// TIA Portal project "ETI C 25" (V15.1)

(* hardware
DEVICE "ET 200SP station_1"  ET 200SP-Station
   slot 0: "Rack_0"  Rack  6ES5 710-8MAx1
   slot 1: "PLC_1"  CPU 1512SP-1 PN  6ES7 512-1DK01-0AB0  V2.6
   slot 2: "DI 16x24VDC ST_1"  DI 16x24VDC ST  6ES7 131-6BH01-0BA0  V0.0
      slot 1: "DI 16x24VDC ST_1"  DI 16x24VDC ST
   slot 3: "DI 16x24VDC ST_2"  DI 16x24VDC ST  6ES7 131-6BH01-0BA0  V0.0
      slot 1: "DI 16x24VDC ST_2"  DI 16x24VDC ST
   slot 4: "DQ 16x24VDC/0.5A ST_1"  DQ 16x24VDC/0.5A ST  6ES7 132-6BH01-0BA0  V0.0
      slot 1: "DQ 16x24VDC/0.5A ST_1"  DQ 16x24VDC/0.5A ST
   slot 5: "AQ 4xU/I ST_1"  AQ 4xU/I ST  6ES7 135-6HD00-0BA1  V1.1
      slot 1: "AQ 4xU/I ST_1"  AQ 4xU/I ST
   slot 6: "Server module_1"  Server module  6ES7 193-6PA00-0AA0  V1.1
      slot 1: "Server module_1"  Server module
   slot 127: "BA 2xRJ45"  BA 2xRJ45  6ES7 193-6AR00-0AA0  V0.0
      slot 32769: "Port_1"  6ES7 193-6AR00-0AA0
      slot 32770: "Port_2"  6ES7 193-6AR00-0AA0
DEVICE "GSD device_1"  GSD.Device.PN
   slot 0: "Rack"  Rack  V1.0
   slot 0: "IOL_I_16_HUB"  IOL_I/O_ 4/ 4 Byte
   slot 0: "mvk1"  55162 MVK DIO12 DIO4/IOL4 M12L 4P  55162  1.08.10
      slot 0: "55162 MVK DIO12 DIO4/IOL4 M12L 4P_1"  55162 MVK DIO12 DIO4/IOL4 M12L 4P
      slot 1: "55162 MVK DIO12 DIO4/IOL4 M12L 4P 1"  55162 MVK DIO12 DIO4/IOL4 M12L 4P
         slot 1: "Port 1"  Port 1
         slot 2: "Port 2"  Port 2
      slot 1: "Device_1"  Device
         slot 0: "Parameter/Diagnostic"  Parameter/Diagnostic
         slot 1: "Digital IO"  Digital IO
      slot 2: "IO-Link master_1"  IO-Link master
   slot 1: "Deactivated"  Deactivated
   slot 2: "Qualifier DI"  Qualifier DI
   slot 2: "FESTO_propocionalniVentil"  IOL_I/O_ 8/ 8 Byte
   slot 3: "Qualifier DO"  Qualifier DO
   slot 3: "SDAT1"  IOL_I_ 2 Byte
   slot 4: "System state"  System state
DEVICE "GSD device_2"  GSD.Device.PN
   slot 0: "Rack"  Rack  V1.0
   slot 0: "IOL_I/O_ 4/ 4 Byte"  IOL_I/O_ 4/ 4 Byte
   slot 0: "mvk2"  55162 MVK DIO12 DIO4/IOL4 M12L 4P  55162  1.08.10
      slot 0: "55162 MVK DIO12 DIO4/IOL4 M12L 4P_1"  55162 MVK DIO12 DIO4/IOL4 M12L 4P
      slot 1: "55162 MVK DIO12 DIO4/IOL4 M12L 4P 2"  55162 MVK DIO12 DIO4/IOL4 M12L 4P
         slot 1: "Port 1"  Port 1
         slot 2: "Port 2"  Port 2
      slot 1: "Device_1"  Device
         slot 0: "Parameter/Diagnostic"  Parameter/Diagnostic
         slot 1: "Digital IO"  Digital IO
      slot 2: "IO-Link master_1"  IO-Link master
   slot 1: "MURR_MVP_2"  IOL_I_ 2 Byte
   slot 2: "Qualifier DI"  Qualifier DI
   slot 2: "IOL_BANNER_LED"  IOL_O_ 4 Byte
   slot 3: "Qualifier DO"  Qualifier DO
   slot 3: "FESTO_SDE1_PRITISK"  IOL_I_ 2 Byte
   slot 4: "System state"  System state
DEVICE "GSD device_3"  GSD.Device.PN
   slot 0: "Rack"  Rack  V1.0
   slot 0: "mvk3"  54504 SOLID67 IOL8 60mm M12L 5P  54504  2.1.1
      slot 0: "DAP"  DAP
      slot 1: "PN-IO"  PN-IO
         slot 1: "Port X01 10/100 MBit/s"  Port X01 10/100 MBit/s
         slot 2: "Port X02 10/100 MBit/s"  Port X02 10/100 MBit/s
      slot 1: "IO-Link Master_1"  IO-Link Master  1.0
         slot 0: "Status/Control Module"  Status/Control Module  1.0
   slot 1: "IFM_VS_temp_pretok"  IO-Link In 4 Bytes
   slot 2: "Digital In (A)/Dig. (B)_1"  Digital In (A)/Dig. (B)
   slot 3: "Digital In (A)/Dig. (B)_2"  Digital In (A)/Dig. (B)
   slot 4: "Digital In (A)/Dig. (B)_3"  Digital In (A)/Dig. (B)
   slot 5: "Digital Out (A)/Dig. (B)"  Digital Out (A)/Dig. (B)
   slot 6: "Digital Out (A)/Dig. (B)_1"  Digital Out (A)/Dig. (B)
   slot 7: "Kamera"  Digital In (A)/Dig. (B)
   slot 8: "FESTO Pnevmatski BLok IO-Link I/O 8/8 Bytes"  IO-Link I/O 8/8 Bytes
DEVICE "GSD device_4"  GSD.Device.PN
   slot 0: "Rack"  Rack  V1.0
   slot 0: "varilnik"  PSS6000 Weld Timer (2-Port)  PSS6000  V1.13.1
      slot 0: "RT"  RT
      slot 1: "Interface"  Interface
         slot 1: "Port 1"  Port 1
         slot 2: "Port 2"  Port 2
   slot 1: "PSI6xxx.780_1"  PSI6xxx.780
      slot 0: "PSI6xxx.780"  PSI6xxx.780
DEVICE "GSD device_7"  GSD.Device.PN
   slot 0: "Rack"  Rack  V1.0
   slot 0: "akd"  AKD-PN-DEVICE  AKD-Pxxxxx-xxPN-xxxx  V00.02
      slot 0: "IDS_SUBMODULE_PARAMDAP"  IDS_SUBMODULE_PARAMDAP
      slot 1: "Interface"  Interface
         slot 1: "Port_1"  Port
   slot 1: "Standard telegram 9_1"  Standard telegram 9  1.0
      slot 0: "Standard telegram 9"  Standard telegram 9
DEVICE "GSD device_5"  GSD.Device.PN
   slot 0: "Rack"  Rack  V1.0
   slot 0: "kroznik"  AKD-PN-DEVICE  AKD-Pxxxxx-xxPN-xxxx  V00.02
      slot 0: "IDS_SUBMODULE_PARAMDAP"  IDS_SUBMODULE_PARAMDAP
      slot 1: "Interface"  Interface
         slot 1: "Port_1"  Port
   slot 1: "Standard telegram 9_1"  Standard telegram 9  1.0
      slot 0: "Standard telegram 9"  Standard telegram 9
DEVICE "GSD device_6"  GSD.Device.PN
   slot 0: "Rack"  Rack  V1.0
   slot 0: "cilinder"  AKD-PN-DEVICE  AKD-Pxxxxx-xxPN-xxxx  V00.02
      slot 0: "IDS_SUBMODULE_PARAMDAP"  IDS_SUBMODULE_PARAMDAP
      slot 1: "Interface"  Interface
         slot 1: "Port_1"  Port
   slot 1: "Standard telegram 9_1"  Standard telegram 9  1.0
      slot 0: "Standard telegram 9"  Standard telegram 9
DEVICE "TP1200 Comfort"  TP1200 Comfort
   slot 0: "TP1200 Comfort"  TP1200 Comfort  6AV2 124-0MC01-0AX0  15.0.0.0
   slot 1: "HMI_RT_6"  TP1200 Comfort  6AV2 124-0MC01-0AX0  15.0.0.0
   slot 5: "TP900 Comfort._CP_1"  PROFINET Interface  15.0.0.0
      slot 1: "PROFINET Interface_1"  PROFINET Interface
         slot 1: "Port_1"  Port
         slot 2: "Port_2"  Port
   slot 7: "TP900 Comfort.I/DP_CP_1"  MPI/DP Interface  15.0.0.0
DEVICE "GSD device_8"  GSD.Device.PN
   slot 0: "Rack"  Rack  V1.0
   slot 0: "dl-pn1"  DL-PN1  DL-PN1  1.00
      slot 0: "DL-PN1"  DL-PN1  1.00
      slot 1: "Interface"  Interface
         slot 1: "Port 1"  Port 1
   slot 1: "DL-PN1_1"  DL-PN1
      slot 0: "DL-PN1 Device"  DL-PN1 Device
   slot 2: "GT2-***_1"  GT2-***
      slot 0: "GT2-***"  GT2-***
   slot 3: "GT2-***_2"  GT2-***
      slot 0: "GT2-***"  GT2-***
*)

// ===== PLC "PLC_1"  CPU 1512SP-1 PN =====

VAR_GLOBAL   // PLC tag table "Default tag table"
   "System_Byte" AT %MB1 : Byte;
   "FirstScan" AT %M1.0 : Bool;
   "DiagStatusUpdate" AT %M1.1 : Bool;
   "AlwaysTRUE" AT %M1.2 : Bool;
   "AlwaysFALSE" AT %M1.3 : Bool;
   "Clock_Byte" AT %MB0 : Byte;
   "Clock_10Hz" AT %M0.0 : Bool;
   "Clock_5Hz" AT %M0.1 : Bool;
   "Clock_2.5Hz" AT %M0.2 : Bool;
   "Clock_2Hz" AT %M0.3 : Bool;
   "Clock_1.25Hz" AT %M0.4 : Bool;
   "Clock_1Hz" AT %M0.5 : Bool;
   "Clock_0.625Hz" AT %M0.6 : Bool;
   "Clock_0.5Hz" AT %M0.7 : Bool;
   "Tag_1" AT %M20.0 : Bool;
   "Tag_2" AT %QD24 : DWord;
   "Tag_3" AT %MD400 : DWord;
   "Tag_4" AT %QD28 : DWord;
   "STOP_SR" AT %M2.0 : Bool;
   "RočnoMerker" AT %M2.2 : Bool;
   "vkloprocno" AT %M2.6 : Bool;
   "RežimDelovanja" AT %MB3 : Byte;
   "BANNER_B3" AT %QB25 : Byte;
   "BANNER_B2" AT %QB26 : Byte;
   "BANNER_B1" AT %QB27 : Byte;
   "BANNER_B0" AT %QB28 : Byte;
   "Tag_5" AT %QW28 : Word;
   "Tag_6" AT %QW25 : Word;
   "Tag_7" AT %QD25 : DWord;
   "STEVEC_KONEC_TRAKA_DOSEZEN" AT %M4.1 : Bool;
   "StatusPrisotnostiTraku" AT %MB5 : Byte;
   "NapakaOdvijanjaTrau" AT %M4.2 : Bool;   // Napaka če se srebrn trak ne odvije
   "NapakaCiscenjaElektrode" AT %M4.3 : Bool;   // Napaka Motorja Čiščenja Traku
   "CiscenjeElektrodeManualOn" AT %M4.4 : Bool;
   "RocniVKlopOdvijanjaTraku" AT %M4.5 : Bool;
   "IzklopStroja" AT %M4.6 : Bool;
   "stevecpreklopov" AT %ID4 : DInt;
   "ZavarjenoSlabiKosi" AT %MD6 : DInt;
   "StartUpBit" AT %M4.7 : Bool;
   "kameratrigger" AT %M10.0 : Bool;
   "ST_IZDELKOV" AT %MD16 : DInt;   // STEVEC KOSOV
END_VAR

VAR_GLOBAL   // PLC tag table "MVK1"
   "MVK_b0" AT %IB20 : Byte;
   "MVK_b1" AT %IB21 : Byte;
   "MVK_b2" AT %IB22 : Byte;
   "MVK_b3" AT %IB23 : Byte;
   "MVK_dw" AT %ID20 : DWord;
   "MVK1_w0" AT %IW20 : Word;
   "ZaporaIzdelka" AT %I20.0 : Bool;   // Y1/1
   "SprositevZaporeIzdelka" AT %I20.1 : Bool;   // Y1/1
   "PrijemaloKontaktaZaprto" AT %I20.2 : Bool;   // Y3/1
   "PrijemaloKontaktaOdprto" AT %I20.3 : Bool;   // Y3/1
   "PozKontaktNaKoncuLetve" AT %I20.4 : Bool;   // Kontakt na koncu letve
   "NC_20.5" AT %I20.5 : Bool;   // NC
   "PozKontaktNaprej" AT %I20.6 : Bool;   // Pozicioniranje pred varjenjem
   "PozKontaktNazaj" AT %I20.7 : Bool;   // Pozicioniranjem pred varjenjem
   "DrzanjeIzmetKontakta" AT %I21.0 : Bool;   // Odpiranje dzanja kontakta nazaj
   "DrzanjeKontakta" AT %I21.1 : Bool;   // Izmet kontakta nazaj
   "IzmetKontaktaNazaj" AT %I21.2 : Bool;   // Izmet vzvoda je v izhodiscu
   "NC_21.3" AT %I21.3 : Bool;   // NC
   "DrcaDobriKosi" AT %I21.4 : Bool;   // Pozicija za dobre kose
   "DrscaSLabiKosi" AT %I21.5 : Bool;   // Pozicija za slabe kose
   "SenzorOdvijanjaCiscenjeElektrode" AT %I21.6 : Bool;   // SenzorCiscenjaElektrode
   "NC_21.7" AT %I21.7 : Bool;
END_VAR

VAR_GLOBAL   // PLC tag table "MVK2"
   "MVK2_b0" AT %IB8 : Byte;
   "MVK2_b1" AT %IB9 : Byte;
   "MVK2_b2" AT %IB10 : Byte;
   "MVK2_b3" AT %IB11 : Byte;
   "MVK2_dw" AT %ID8 : DWord;
   "MVK2_w0" AT %IW8 : Word;
   "MVK2_w1" AT %IW10 : Word;
   "KAMERA_FEEDBACK" AT %I8.0 : Bool;
   "NC_8.1" AT %I8.1 : Bool;
   "NC_8.2" AT %I8.2 : Bool;
   "NC_8.3" AT %I8.3 : Bool;
   "SenzorStartOdvijanje" AT %I8.4 : Bool;   // Senzor za začetek odvijanja koluta
   "SenzorKoluta" AT %I8.5 : Bool;   // Senzor za detekcijo odvijanja koluta
   "PrisotnostTraka" AT %I8.6 : Bool;
   "NC_8.7" AT %I8.7 : Bool;
   "RazsvetljavaLevo" AT %Q20.0 : Bool;
   "RazsvetljavaDesno" AT %Q20.1 : Bool;
   "NC_Q20.2" AT %Q20.2 : Bool;
   "NC_Q20.3" AT %Q20.3 : Bool;
   "NC_Q20.4" AT %Q20.4 : Bool;
   "NC_Q20.5" AT %Q20.5 : Bool;
   "NC_Q20.6" AT %Q20.6 : Bool;
   "NC_Q20.7" AT %Q20.7 : Bool;
END_VAR

VAR_GLOBAL   // PLC tag table "SDAT"
   "I_SDAT1" AT %IW32 : Word;   // Y2/1
   "I_SDAT2" AT %IW34 : Word;   // Y1/2
END_VAR

VAR_GLOBAL   // PLC tag table "MURR IOL M"
   "MURR_IOL1_DO" AT %QB0 : Byte;
   "SoftStart" AT %Q0.0 : Bool;   // SOFTSTART - vklop pnevmatike
   "MURR_IOL1_DO.1" AT %Q0.1 : Bool;
   "MURR_IOL1_DO.2" AT %Q0.2 : Bool;   // Napajanje IOL power supply
   "MURR_IOL1_DO.3" AT %Q0.3 : Bool;
   "MURR_IOL1_DO.4" AT %Q0.4 : Bool;
   "MURR_IOL1_DO.5" AT %Q0.5 : Bool;
   "MURR_IOL1_DO.6" AT %Q0.6 : Bool;
   "MURR_IOL1_DO.7" AT %Q0.7 : Bool;
   "MURR_IOL2_DO" AT %QB2 : Byte;
   "MURR_IOL2_DO.0" AT %Q2.0 : Bool;
   "MURR_IOL2_DO.1" AT %Q2.1 : Bool;
   "MURR_IOL2_DO.2" AT %Q2.2 : Bool;
   "MURR_IOL2_DO.3" AT %Q2.3 : Bool;
   "MURR_IOL2_DO.4" AT %Q2.4 : Bool;
   "MURR_IOL2_DO.5" AT %Q2.5 : Bool;
   "MURR_IOL2_DO.6" AT %Q2.6 : Bool;
   "MURR_IOL2_DO.7" AT %Q2.7 : Bool;
   "FESTO_pritisk" AT %IW52 : Word;
   "PropocionalniVentilSet" AT %QW32 : Word;
   "PropocionalniVentilTrenutna" AT %IW44 : Word;
END_VAR

VAR_GLOBAL   // PLC tag table "FESTO"
   "FESTO_W0" AT %QW44 : Word;
   "FESTO_W1" AT %QW46 : Word;
   "FESTO_W2" AT %QW48 : Word;
   "FESTO_W3" AT %QW50 : Word;
   "1Y1_OdklepZapore" AT %Q44.0 : Bool;
   "Y2/1_NalaganjeNaprej" AT %Q44.2 : Bool;
   "Y2/1_NalaganjeNazanj" AT %Q44.3 : Bool;
   "Y3/1_PrijemaloKontaktaOdpri" AT %Q44.4 : Bool;
   "Y3/1_NC" AT %Q44.5 : Bool;
   "Y1/3_OdmičniCilinderKonusa" AT %Q45.0 : Bool;
   "Y1/3_NC" AT %Q45.1 : Bool;
   "Y2/3_PozicioniranjeKontaktovNazaj" AT %Q45.2 : Bool;
   "Y2/3_PozicioniranjeKontaktovNaprej" AT %Q45.3 : Bool;
   "Y3/3_OdpiranjeDržalaKomada" AT %Q45.4 : Bool;
   "Y3/3_NC" AT %Q45.5 : Bool;
   "Y4/3_OdpiranjeIzmetaKontakta" AT %Q45.6 : Bool;
   "Y4/3_NC" AT %Q45.7 : Bool;
   "Y5/3_IzmetKomadov" AT %Q46.0 : Bool;
   "Y5/3_NC" AT %Q46.1 : Bool;
   "Y6/3_LoputaDobri" AT %Q46.2 : Bool;
   "Y6/3_LoputaSlabi" AT %Q46.3 : Bool;
   "Y1/4_odmičniCilinderVarjenje_GOR" AT %Q46.4 : Bool;
   "Y1/4_odmičniCilinderVarjenjeDOL" AT %Q46.5 : Bool;
   "ČiščenjeElektrode_ON" AT %Q46.6 : Bool;
   "ČiščenjeElektrode_OFF" AT %Q46.7 : Bool;
   "PihanjeLinearniVibrator" AT %Q47.0 : Bool;
   "NC" AT %Q47.1 : Bool;
   "Y2/1_dovajanjePlosciceNazaj" AT %Q44.6 : Bool;
   "Y2_1_dovajanjePlosciceNaprej" AT %Q44.7 : Bool;
   "1Y1_zaklep_NC" AT %Q44.1 : Bool;
END_VAR

VAR_GLOBAL   // PLC tag table "MVK3"
   "MVK3_b0" AT %QB40 : Byte;
   "MVK3_b1" AT %QB41 : Byte;
   "MVK3_b2" AT %QB42 : Byte;
   "MVK3_b4" AT %QB43 : Byte;
   "MVK3_O_X1_P4" AT %Q40.0 : Bool;
   "MVK3_O_X1_P2" AT %Q40.1 : Bool;
   "MVK3_O_X2_P4" AT %Q40.2 : Bool;
   "MVK3_O_X2_P2" AT %Q40.3 : Bool;
   "MVK3_O_X3_P4" AT %Q40.4 : Bool;
   "MVK3_O_X3_P2" AT %Q40.5 : Bool;
   "MVK3_O_X4_P4" AT %Q40.6 : Bool;
   "MVK3_O_X4_P2" AT %Q40.7 : Bool;
   "MVK3_O_X5_P4_NC" AT %Q41.0 : Bool;   // X5,P4 - PIN 4 NC
   "RazsvetljavaSpredaj" AT %Q41.1 : Bool;   // 5404 IOL X5, P2 - MASTER - PIN2/5 - razsvetljava LED SPREDAJ
   "bTrigOptoEnginering" AT %Q41.2 : Bool;   // X6, P4 : triger za led
   "bVccOptoEngineering" AT %Q41.3 : Bool;   // X6, P2 : Vklop napajanja
   "MVK3_O_b1.4" AT %Q41.4 : Bool;   // X7, P4
   "MVK3_O_b1.5" AT %Q41.5 : Bool;   // X7, P2
   "MVK3_O_b1.6" AT %Q41.6 : Bool;   // X8, P4
   "MVK3_O_b1.7" AT %Q41.7 : Bool;   // X8,P2
   "MVK3_O_b2.0" AT %Q42.0 : Bool;
   "MVK3_O_b2.1" AT %Q42.1 : Bool;
   "MVK3_O_b2.2" AT %Q42.2 : Bool;
   "MVK3_O_b2.3" AT %Q42.3 : Bool;
   "MVK3_O_b2.4" AT %Q42.4 : Bool;
   "MVK3_O_b2.5" AT %Q42.5 : Bool;
   "MVK3_O_b2.6" AT %Q42.6 : Bool;
   "MVK3_O_b2.7" AT %Q42.7 : Bool;
   "MVK3_O_b3.0" AT %Q43.0 : Bool;
   "MVK3_O_b3.1" AT %Q43.1 : Bool;
   "MVK3_O_b3.2" AT %Q43.2 : Bool;
   "MVK3_O_b3.3" AT %Q43.3 : Bool;
   "MVK3_O_b3.4" AT %Q43.4 : Bool;
   "MVK3_O_b3.5" AT %Q43.5 : Bool;
   "MVK3_O_b3.6" AT %Q43.6 : Bool;
   "MVK3_O_b3.7" AT %Q43.7 : Bool;
   "IOL_IFM_SV" AT %ID36 : DWord;
   "MVK3_I_b0" AT %IB54 : Byte;
   "MVK3_I_b1" AT %IB55 : Byte;
   "MVK3_I_b2" AT %IB56 : Byte;
   "MVK3_I_b3" AT %IB57 : Byte;
END_VAR

VAR_GLOBAL   // PLC tag table "PLC_IO"
   "PLC_I_W0" AT %IW0 : Word;
   "PLCI_W2" AT %IW2 : Word;
   "PLC_I0.0" AT %I0.0 : Bool;   // DC OK
   "IzklopVsiliBtnPanel" AT %I0.1 : Bool;
   "VarmostZavese" AT %I0.2 : Bool;   // VarnostneZavese [1-ok, 0, nok]
   "PremostitevVarnostiBtnPanel" AT %I0.3 : Bool;
   "PrisotnostIzmetaIzdelka" AT %I0.4 : Bool;   // Senzor Izmeta na koncu traku
   "PLC_I0.5" AT %I0.5 : Bool;
   "PLC_I0.6" AT %I0.6 : Bool;
   "PLC_I0.7" AT %I0.7 : Bool;
   "PLC_I1.0" AT %I1.0 : Bool;
   "PLC_I1.1" AT %I1.1 : Bool;
   "RežimRočno" AT %I1.2 : Bool;
   "RežimAvtomatsko" AT %I1.3 : Bool;
   "StartCiklaBtnPanel" AT %I1.4 : Bool;
   "StopCiklaBtnPanel" AT %I1.5 : Bool;
   "ResetNapake" AT %I1.6 : Bool;
   "VklopKrmiljaBtnPanel" AT %I1.7 : Bool;
   "VKlopvarnostnegaModulaIVS" AT %QW4 : Word;
   "VklopVarnosnegaModula" AT %Q4.0 : Bool;
   "VklopZaves" AT %Q4.1 : Bool;
   "NightShift" AT %Q4.2 : Bool;
   "AKD_sprostitevZavore" AT %Q4.3 : Bool;
   "PLC_Q4.4" AT %Q4.4 : Bool;
   "PLC_Q4.5" AT %Q4.5 : Bool;
   "PLC_Q4.6" AT %Q4.6 : Bool;
   "VentilVode" AT %Q4.7 : Bool;
   "PLC_Q5.0" AT %Q5.0 : Bool;
   "MotorOdvijanjeTraku" AT %Q5.1 : Bool;
   "MotorČiščenjeElektrode" AT %Q5.2 : Bool;
   "LED_RUN" AT %Q5.3 : Bool;
   "LED_ERROR" AT %Q5.4 : Bool;
   "AKD_HW_ENABLE" AT %Q5.5 : Bool;
   "TekociTrakVklop" AT %Q5.6 : Bool;
   "PolnjenjeSkatle1" AT %Q5.7 : Bool;
   "+" AT %I2.0 : Bool;
   "-" AT %I2.1 : Bool;
   "i2.0_b2" AT %I2.2 : Bool;
   "i2.0_b3" AT %I2.3 : Bool;
   "i2.0_b4" AT %I2.4 : Bool;
   "i2.0_b5" AT %I2.5 : Bool;
   "i2.0_b6" AT %I2.6 : Bool;
   "i2.0_b7" AT %I2.7 : Bool;
   "i2.0_b8" AT %I3.0 : Bool;
   "i2.0_b9" AT %I3.1 : Bool;
   "i2.0_b10" AT %I3.2 : Bool;
   "i2.0_b11" AT %I3.3 : Bool;
   "i2.0_b12" AT %I3.4 : Bool;
   "i2.0_b13" AT %I3.5 : Bool;
   "i2.0_b14" AT %I3.6 : Bool;
END_VAR

VAR_GLOBAL   // PLC tag table "VARJENJE"
   "Varjenje_QB0" AT %QB52 : Byte;
   "Varjenje_QB1" AT %QB53 : Byte;
   "Varjanje_IB0" AT %IB66 : Byte;
   "Varjenje_IB0" AT %IB67 : Byte;
   "ValidSpotSelection" AT %Q52.0 : Bool;
   "Varjenje_Qb0.1" AT %Q52.1 : Bool;
   "Start" AT %Q52.2 : Bool;
   "GeneralFaultReset" AT %Q52.3 : Bool;
   "ResetWithEOS" AT %Q52.4 : Bool;
   "ResetWithReweld" AT %Q52.5 : Bool;
   "Varjenje_Qb0.6" AT %Q52.6 : Bool;
   "Varjenje_Qb0.7" AT %Q52.7 : Bool;
   "ExternalWeldOn" AT %Q53.0 : Bool;
   "Varjenje_Qb1.1" AT %Q53.1 : Bool;
   "Varjenje_Qb1.2" AT %Q53.2 : Bool;
   "Varjenje_Qb1.3" AT %Q53.3 : Bool;
   "Varjenje_Qb1.4" AT %Q53.4 : Bool;
   "Varjenje_Qb1.5" AT %Q53.5 : Bool;
   "Varjenje_Qb1.6" AT %Q53.6 : Bool;
   "Varjenje_Qb1.7" AT %Q53.7 : Bool;
   "Varjenje_Qb2.0" AT %Q54.0 : Bool;
   "Varjenje_Qb2.1" AT %Q54.1 : Bool;
   "Varjenje_Qb2.2" AT %Q54.2 : Bool;
   "Varjenje_Qb2.3" AT %Q54.3 : Bool;
   "Varjenje_Qb2.4" AT %Q54.4 : Bool;
   "Varjenje_Qb2.5" AT %Q54.5 : Bool;
   "Varjenje_Qb2.7" AT %Q54.7 : Bool;
   "Varjenje_Qb2.8" AT %Q55.0 : Bool;
   "Varjenje_Qb2.9" AT %Q55.1 : Bool;
   "Varjenje_Qb2.10" AT %Q55.2 : Bool;
   "Varjenje_Qb2.11" AT %Q55.3 : Bool;
   "Varjenje_Qb2.12" AT %Q55.4 : Bool;
   "SpotSelection" AT %QB60 : Byte;
   "SpotSelectionTakeOver" AT %I66.0 : Bool;   // Program izbran
   "Varjenje_Ib0.1" AT %I66.1 : Bool;
   "EndOfSequency_WC" AT %I66.2 : Bool;   // Konec varjenja
   "TimerReady" AT %I66.3 : Bool;   // Varilnik pripravljen
   "WeldFault" AT %I66.4 : Bool;   // Napaka varjenja
   "Varjenje_Ib0.5" AT %I66.5 : Bool;
   "Varjenje_Ib0.6" AT %I66.6 : Bool;
   "Varjenje_Ib0.7" AT %I66.7 : Bool;
   "FiringEnable" AT %I67.0 : Bool;   // Varjenje Vključeno
   "Varjenje_Ib2.1" AT %I67.1 : Bool;
   "Varjenje_Ib2.2" AT %I67.2 : Bool;
   "Varjenje_Ib2.3" AT %I67.3 : Bool;
   "Varjenje_Ib2.4" AT %I67.4 : Bool;
   "Varjenje_Ib2.5" AT %I68.0 : Bool;
   "Varjenje_Ib2.6" AT %I68.1 : Bool;
   "Varjenje_Ib2.7" AT %I68.2 : Bool;
   "Varjenje_Ib2.8" AT %I68.3 : Bool;
   "Varjenje_Ib2.9" AT %I68.4 : Bool;
   "Varjenje_Ib2.10" AT %I68.5 : Bool;
   "StatusCode" AT %IB82 : Byte;   // Status
   "Status_b0" AT %IB80 : Byte;
   "Status_b1" AT %IB83 : Byte;
   "Varjenje_Qb2.6" AT %Q54.6 : Bool;
END_VAR

VAR_GLOBAL   // PLC tag table "AKD_elektroda"
   "PogojZaservoOn" AT %M2.1 : Bool;
   "tipka+" AT %M2.3 : Bool;
   "tipka-" AT %M2.4 : Bool;
   "ElektrodaSiemensToAkd" AT %Q400.0 : "SIEMENS_TO_AKD";
   "ElektrodaAkdToSiemens" AT %I400.0 : "AKD_TO_SIEMENS";
   "onemogoci" AT %M2.7 : Bool;
   "enable" AT %M4.0 : Bool;
   "STEVEC_KOSOV" AT %C0 : Counter;
   "manualCameraTrig" AT %M10.1 : Bool;   // trig kamera
   "MotorCiscenjeElektrodeCOunter" AT %MD12 : DInt;   // Stevec
   "prisotnostizmetaarker" AT %M10.2 : Bool;   // Merker za R edge - izmeta kontakta - senzor
END_VAR

VAR_GLOBAL   // PLC tag table "AKD_kroznik"
   "KroznikSiemensToAkd" AT %Q98.0 : "SIEMENS_TO_AKD";
   "KroznikAkdToSiemens" AT %I98.0 : "AKD_TO_SIEMENS";
   "servpen" AT %M2.5 : Bool;
END_VAR

VAR_GLOBAL   // PLC tag table "AKD_REZANJEPODAJANJE"
   "rezanjepodajanjeSiemenstoAKD" AT %I108.0 : "AKD_TO_SIEMENS";
   "rezanjepodajanje_SiemensToAKD" AT %Q118.0 : "SIEMENS_TO_AKD";
END_VAR

VAR_GLOBAL   // PLC tag table "KEYENCE"
   "Keyence_OdmičniCilinderKonusa" AT %ID137 : DInt;   // Cilinder odmika mize
   "Keyence_OdmičniCilinderVarjenja" AT %ID144 : DInt;   // Cilinder odmika varjenja
END_VAR

TYPE "UDT_MVK1"
   STRUCT
      "1Y1" : Struct   // VKLOP/IZKLOP zapore na LIN vibratorju
         B1 : Bool;   // POZ Zaklep linearnega vibratorja
         B2 : Bool;   // POZ Odklep linearnega vibratorja
      END_STRUCT;
      "Y3/1" : Struct   // Prijemalo kontakta
         B1 : Bool;   // POZ Prijemalo zaprto
         B2 : Bool;   // POZ Prijemalo odprto
      END_STRUCT;
      B_kontaktnaKoncuLetve : Struct   // Detekcija kontakta na letvi
         B1 : Bool;   // POZ kontakt na koncu letve
         NC : Bool;
      END_STRUCT;
      "Y2/3" : Struct   // Pozicioniranje kontakta
         B1 : Bool;   // POZ kontakta naprej
         B2 : Bool;   // POZ Prijemalo odprto
      END_STRUCT;
      "Y3/3" : Struct   // Držanje kontakta v mizi
         B1 : Bool;   // POZ držanje kontakta odprto
      END_STRUCT;
      "Y4/3" : Struct   // Odpiranje izmeta konkta
         B1 : Bool;   // POZ izmet kontakta odprt
      END_STRUCT;
      "Y5/3" : Struct   // Izmet kontakta
         B1 : Bool;   // POZ izmet kontakta nazaj
      END_STRUCT;
      "Y6/3" : Struct   // Drča dobri/slabi kosi
         B1 : Bool;   // POZ dobri kosi
         B2 : Bool;   // POZ slabi kosi
      END_STRUCT;
      KonrolaIzmeta : Struct   // kontrola izmeta
         IzmetOK : Bool;   // Senzor preleta izmeta
         NC : Bool;
      END_STRUCT;
   END_STRUCT;
END_TYPE

TYPE "SIEMENS_TO_AKD"
   STRUCT
      PODATKI : Struct
         oBit8_jogOn : Bool;   // b0
         oBit9_jog2On : Bool;   // 1
         ControlByPLC : Bool;   // 2
         StartHomming : Bool;   // 3
         NC_B0_b4 : Bool;   // 4
         NC_B0_b5 : Bool;   // 5
         NC_B0_b6 : Bool;   // 6
         NC_B0_b7 : Bool;   // 7
         SwtichOn : Bool;   // 0
         NoCoastStop : Bool;   // 1
         NoQuickStop : Bool;   // 2
         EnableOperation : Bool;   // 3
         EnableRampGen : Bool;   // 4
         UnfreezeRamp : Bool;   // 5
         EnableSetPoint : Bool;   // 6
         FaultAckt : Bool;   // 7 1
         SATANW : Int;   // 0- 26 2-3
         byte4 : Byte;   // 4
         byte5 : Byte;   // 5
         MDI_TARPOS : DInt;   // 6 7 8 9
         MDI_VELOCITY : DInt;   // 10 11 12 13
         b14 : DInt;   // 14
         "15" : DInt;   // 15
         b16 : DInt;   // 16
         b17 : DInt;   // 17
         MDI_MOD : DInt;   // 18,19
      END_STRUCT;
   END_STRUCT;
END_TYPE

TYPE "AKD_TO_SIEMENS"
   STRUCT
      PODATKI_TO_SIEMENS : Struct
         ErrInRange : Bool;
         ContrReqByMass : Bool;
         TargetPosreached : Bool;
         HomePosSet : Bool;
         TravesingTaskAck : Bool;
         DriveStopen : Bool;
         MotionTaskActive : Bool;
         "i_b0.7" : Bool;
         ReadyToSwitch : Bool;
         ReadyToOperate : Bool;
         OperationENabled : Bool;
         FaultPresent : Bool;
         CoastStopNotAct : Bool;
         QuickStopNotAct : Bool;
         SwitchOnInhibiited : Bool;
         WarningPreent : Bool;
         AKTSATZ : Word;
         ZSW2 : Word;
         ActualPos : DWord;
      END_STRUCT;
   END_STRUCT;
END_TYPE

TYPE "PDT_AKD"
   STRUCT
      PODATKI : Struct
         AKDenable : Bool;
         NastavitevHitrosti : Int := 60;
         NastavitevPozicije : DInt := 12;
         TrenutnaPozicija : DInt;
         ServoGo : Bool;
         StartHomming : Bool;
      END_STRUCT;
   END_STRUCT;
END_TYPE

TYPE "BOSH"
   STRUCT
      PDT_BOSH_STATUS : Struct
         OK : UInt := 0;
         IZKLOP_V_SILI : UInt := 80;
         WELD_WITHOUD_COMMAND : UInt := 81;
         MEMMORY_DELETED : UInt := 85;
         DATA_DOWNLOAD_ACTIVE : UInt := 86;
         NO_WELDING_PROGRAM : UInt := 87;
         HARDWARE_FAULT : UInt := 88;
         "I/O_BUS_FAULT" : UInt := 89;
         HWAVE_MONITORING : UInt := 90;
         MAIN_SWITCH_TRIPPED : UInt := 91;
         EXTERNAL_TEMEPERATURE_TO_HIGH : UInt := 92;
         SYC_ERROR : UInt := 93;
         START_INHIBITED : UInt := 94;
         PROGRAM_PARITY_ERROR : UInt := 95;
         PROGRAMED_VALUE_TO_LARGE : UInt := 98;
         WELD_PROCESS_ERROR : UInt := 99;
         SUPPLY_VOLTAGE_VAULT : UInt := 100;
         MAX_HEAT_SINK_TEMP : UInt := 160;
         TRANSFORMER_TEMP_TO_HIGH : UInt := 164;
         HARDWARE_FAULT_DRIVE_MODULE : UInt := 165;
      END_STRUCT;
   END_STRUCT;
END_TYPE

DATA_BLOCK "SDAT1"   // DB1
{ S7_Optimized_Access := 'TRUE' }
VERSION : 0.1
// stored: InstanceOfName FB_IOL_SDAT
"FB_IOL_SDAT"
BEGIN
END_DATA_BLOCK

DATA_BLOCK "SDAT2"   // DB2
{ S7_Optimized_Access := 'TRUE' }
VERSION : 0.1
// stored: InstanceOfName FB_IOL_SDAT
"FB_IOL_SDAT"
BEGIN
END_DATA_BLOCK

DATA_BLOCK "FB_MVK1_DB"   // DB3
{ S7_Optimized_Access := 'TRUE' }
VERSION : 0.1
// stored: InstanceOfName FB_MVK1
"FB_MVK1"
BEGIN
END_DATA_BLOCK

DATA_BLOCK "FB_IOL_IFM_SV_DB"   // DB4
{ S7_Optimized_Access := 'TRUE' }
VERSION : 0.1
// stored: InstanceOfName FB_IOL_IFM_SV
"FB_IOL_IFM_SV"
BEGIN
END_DATA_BLOCK

DATA_BLOCK "FB_FESTO_VPPM_DB"   // DB5
{ S7_Optimized_Access := 'TRUE' }
VERSION : 0.1
// stored: InstanceOfName FB_FESTO_VPPM
"FB_FESTO_VPPM"
BEGIN
END_DATA_BLOCK

DATA_BLOCK "FB_GL_PROGRAM_DB"   // DB6
{ S7_Optimized_Access := 'TRUE' }
VERSION : 0.1
// stored: InstanceOfName FB_GL_PROGRAM
"FB_GL_PROGRAM"
BEGIN
END_DATA_BLOCK

DATA_BLOCK "FB_AKD_Kroznik"   // DB8
{ S7_Optimized_Access := 'TRUE' }
VERSION : 0.1
// stored: InstanceOfName FB_AKD
"FB_AKD"
BEGIN
END_DATA_BLOCK

DATA_BLOCK "FB_AKD_REZANJEPODAJANJE"   // DB9
{ S7_Optimized_Access := 'TRUE' }
VERSION : 0.1
// stored: InstanceOfName FB_AKD
"FB_AKD"
BEGIN
END_DATA_BLOCK

DATA_BLOCK "db_AKD"   // DB10
{ S7_Optimized_Access := 'TRUE' }
VERSION : 0.1
   VAR RETAIN
      REZANJEPODAJANJE : Struct
         PODATKI : Struct
            AKDenable : Bool;
            NastavitevHItrosti : Int := 60;
            NastavitevPozicije : Int := 12;
            NastavitevPrograma : Struct
               "Položaj rezanja" : Word := 16#00_00;
               "Položaj podajanja" : Word := 16#00_01;
               IzbranProgram : Word;
            END_STRUCT;
            ServoGO : Bool;
            TrenutnaPozicija : DInt;
            Podano : Bool;
            Odrezano : Bool;
            ZahtevaPoPodajanju : Bool;
            ZahtevaPoRezanju : Bool;
            PloscicaOdrezana : Bool;
            merkerji : Array[0..1] of Bool;
            kokrak : UInt;
            vPODAJANJU : Bool;
            VrEZANJU : Bool;
         END_STRUCT;
      END_STRUCT;
      ELEKTRODA : "PDT_AKD";
      KROZNIK : "PDT_AKD";
   END_VAR
BEGIN
END_DATA_BLOCK

DATA_BLOCK "dbAreaPointer"   // DB11
{ S7_Optimized_Access := 'FALSE' }
VERSION : 0.1
   VAR
      Coordination : Array[0..15] of Bool;
      "Date/Time" : Array[0..5] of Word;
      JobMailbox : Array[0..3] of Word;
      HMIscreenNum : Array[0..4] of Word;
   END_VAR
BEGIN
END_DATA_BLOCK

DATA_BLOCK "FB_STARTUP_DB"   // DB12
{ S7_Optimized_Access := 'TRUE' }
VERSION : 0.1
// stored: InstanceOfName FB_STARTUP
"FB_STARTUP"
BEGIN
END_DATA_BLOCK

DATA_BLOCK "FB_FESTO_SDE1_DB"   // DB13
{ S7_Optimized_Access := 'TRUE' }
VERSION : 0.1
// stored: InstanceOfName FB_FESTO_SDE1
"FB_FESTO_SDE1"
BEGIN
END_DATA_BLOCK

DATA_BLOCK "FB_Lin_FESTO_PNEVMATIKA_PRITISK"   // DB14
{ S7_Optimized_Access := 'TRUE' }
VERSION : 0.1
// stored: InstanceOfName FB_Lin_fun
"FB_Lin_fun"
BEGIN
END_DATA_BLOCK

DATA_BLOCK "DB_HMI"   // DB15
{ S7_Optimized_Access := 'TRUE' }
VERSION : 0.1
   VAR RETAIN
      PREKLOP_HMI : Struct
         merkers : Array[0..10] of Bool;
         HMI_AVTO_nr : Int := 18;   // Št. ekrana v avt. načinu
         HMI_ROČNO_nr : Int := 5;   // št. ekrana v ročnem načinu
      END_STRUCT;
   END_VAR
   VAR
      "ROČNI NAČIN" : Struct
         izbraniCilinder : Int := 220;
      END_STRUCT;
   END_VAR
   VAR RETAIN
      SDAT1 : Struct   // Nalaganje izdelka
         PozPobiranje : Real := 77.7;   // POZ pobiranja komada
         PozNalaganje : Real := 10.9;   // POZ nalaganja komada
      END_STRUCT;
      SDAT2 : Struct   // Nalaganje ploščice
         PozPobiranjePloscice : Real := 70.0;   // POZ pobiranja ploščice
         PozNalaganjePloscice : Real := 11.5;   // POZ nalaganja ploščice
      END_STRUCT;
      Varjenje : Struct
         ResetWithWC : Bool := FALSE;
         ResetWithWeld : Bool := FALSE;
      END_STRUCT;
      TekočiTrak : Struct
         btnResetSkatle1 : Bool := FALSE;
         btnResetSKatle2 : Bool := FALSE;
      END_STRUCT;
      Kroznik : Struct
         bStartHomming : Bool := FALSE;
      END_STRUCT;
      HMI_izpisNapak : Struct
         w_trenutnaNapak : WString;
      END_STRUCT;
      ČiščenjeElektrode : Struct
         ZeljenoStevilo : UInt;
      END_STRUCT;
   END_VAR
BEGIN
   PREKLOP_HMI.merkers[0] := FALSE;   // P merker preklop ročno
   PREKLOP_HMI.merkers[1] := FALSE;   // P merker preklop avtomatsko
   PREKLOP_HMI.merkers[2] := FALSE;
   PREKLOP_HMI.merkers[3] := FALSE;
   PREKLOP_HMI.merkers[4] := FALSE;
   PREKLOP_HMI.merkers[5] := FALSE;
   PREKLOP_HMI.merkers[6] := FALSE;
   PREKLOP_HMI.merkers[7] := FALSE;
   PREKLOP_HMI.merkers[8] := FALSE;
   PREKLOP_HMI.merkers[9] := FALSE;
   PREKLOP_HMI.merkers[10] := FALSE;
END_DATA_BLOCK

DATA_BLOCK "FB_ROČNO_VODENJE_DB"   // DB16
{ S7_Optimized_Access := 'TRUE' }
VERSION : 0.1
// stored: InstanceOfName FB_ROČNO_VODENJE
"FB_ROČNO_VODENJE"
BEGIN
END_DATA_BLOCK

DATA_BLOCK "DB_UDP_COMM"   // DB17
{ S7_Optimized_Access := 'FALSE' }
VERSION : 0.1
   VAR
      PLC_TO_PC : Struct
         PC_addr : TADDR_Param;
         DATA : Array[0..1023] of Char;
         TON_COM_REQ : Bool := FALSE;
         TDIS_COM_REQ : Bool := FALSE;
         TCON_COM_REQ : Bool := FALSE;
         TCON_DB : Struct
            done : Bool := FALSE;
            busy : Bool := FALSE;
            error : Bool := FALSE;
            status : Word := 16#0000;
            con_succ : Bool := FALSE;
         END_STRUCT;
         TUSEND_DB : Struct
            done : Bool := FALSE;
            busy : Bool := FALSE;
            error : Bool := FALSE;
            status : Word := 16#7000;
            TUSEND_REQ : Bool := FALSE;
            SendSucess : Bool := TRUE;
         END_STRUCT;
         TurnOffPC : Bool := FALSE;
         FirstRun : Bool := TRUE;
      END_STRUCT;
      TC_ON_COMM_DATA : Struct
         REQ : Bool := TRUE;
         ID : Bool := FALSE;
         DONE : Bool := FALSE;
         BUSY : Bool := FALSE;
         ERROR : Bool := FALSE;
         STATUS : Word := 16#7000;
      END_STRUCT;
      ConnectionEstablish : Bool := FALSE;
      FirstRun : Bool := FALSE;
   END_VAR
BEGIN
   PLC_TO_PC.PC_addr.REM_IP_ADDR[1] := 192;
   PLC_TO_PC.PC_addr.REM_IP_ADDR[2] := 168;
   PLC_TO_PC.PC_addr.REM_IP_ADDR[3] := 0;
   PLC_TO_PC.PC_addr.REM_IP_ADDR[4] := 200;
   PLC_TO_PC.PC_addr.REM_PORT_NR := 5000;
   PLC_TO_PC.DATA[1] := '$02';
   PLC_TO_PC.DATA[2] := '$01';
   PLC_TO_PC.DATA[3] := '7';
   PLC_TO_PC.DATA[4] := 'B';
   PLC_TO_PC.DATA[5] := '$R';
   PLC_TO_PC.DATA[6] := '$L';
   PLC_TO_PC.PC_addr.RESERVED := 16#0000;
   PLC_TO_PC.DATA[0] := '1';
   PLC_TO_PC.DATA[7] := ' ';
   PLC_TO_PC.DATA[8] := ' ';
   PLC_TO_PC.DATA[9] := ' ';
   PLC_TO_PC.DATA[10] := ' ';
   PLC_TO_PC.DATA[11] := ' ';
   PLC_TO_PC.DATA[12] := ' ';
   PLC_TO_PC.DATA[13] := ' ';
   PLC_TO_PC.DATA[14] := ' ';
   PLC_TO_PC.DATA[15] := ' ';
   PLC_TO_PC.DATA[16] := ' ';
   PLC_TO_PC.DATA[17] := ' ';
   PLC_TO_PC.DATA[18] := ' ';
   PLC_TO_PC.DATA[19] := ' ';
   PLC_TO_PC.DATA[20] := ' ';
   PLC_TO_PC.DATA[21] := ' ';
   PLC_TO_PC.DATA[22] := ' ';
   PLC_TO_PC.DATA[23] := ' ';
   PLC_TO_PC.DATA[24] := ' ';
   PLC_TO_PC.DATA[25] := ' ';
   PLC_TO_PC.DATA[26] := ' ';
   PLC_TO_PC.DATA[27] := ' ';
   PLC_TO_PC.DATA[28] := ' ';
   PLC_TO_PC.DATA[29] := ' ';
   PLC_TO_PC.DATA[30] := ' ';
   PLC_TO_PC.DATA[31] := ' ';
   PLC_TO_PC.DATA[32] := ' ';
   PLC_TO_PC.DATA[33] := ' ';
   PLC_TO_PC.DATA[34] := ' ';
   PLC_TO_PC.DATA[35] := ' ';
   PLC_TO_PC.DATA[36] := ' ';
   PLC_TO_PC.DATA[37] := ' ';
   PLC_TO_PC.DATA[38] := ' ';
   PLC_TO_PC.DATA[39] := ' ';
   PLC_TO_PC.DATA[40] := ' ';
   PLC_TO_PC.DATA[41] := ' ';
   PLC_TO_PC.DATA[42] := ' ';
   PLC_TO_PC.DATA[43] := ' ';
   PLC_TO_PC.DATA[44] := ' ';
   PLC_TO_PC.DATA[45] := ' ';
   PLC_TO_PC.DATA[46] := ' ';
   PLC_TO_PC.DATA[47] := ' ';
   PLC_TO_PC.DATA[48] := ' ';
   PLC_TO_PC.DATA[49] := ' ';
   PLC_TO_PC.DATA[50] := ' ';
   PLC_TO_PC.DATA[51] := ' ';
   PLC_TO_PC.DATA[52] := ' ';
   PLC_TO_PC.DATA[53] := ' ';
   PLC_TO_PC.DATA[54] := ' ';
   PLC_TO_PC.DATA[55] := ' ';
   PLC_TO_PC.DATA[56] := ' ';
   PLC_TO_PC.DATA[57] := ' ';
   PLC_TO_PC.DATA[58] := ' ';
   PLC_TO_PC.DATA[59] := ' ';
   PLC_TO_PC.DATA[60] := ' ';
   PLC_TO_PC.DATA[61] := ' ';
   PLC_TO_PC.DATA[62] := ' ';
   PLC_TO_PC.DATA[63] := ' ';
   PLC_TO_PC.DATA[64] := ' ';
   PLC_TO_PC.DATA[65] := ' ';
   PLC_TO_PC.DATA[66] := ' ';
   PLC_TO_PC.DATA[67] := ' ';
   PLC_TO_PC.DATA[68] := ' ';
   PLC_TO_PC.DATA[69] := ' ';
   PLC_TO_PC.DATA[70] := ' ';
   PLC_TO_PC.DATA[71] := ' ';
   PLC_TO_PC.DATA[72] := ' ';
   PLC_TO_PC.DATA[73] := ' ';
   PLC_TO_PC.DATA[74] := ' ';
   PLC_TO_PC.DATA[75] := ' ';
   PLC_TO_PC.DATA[76] := ' ';
   PLC_TO_PC.DATA[77] := ' ';
   PLC_TO_PC.DATA[78] := ' ';
   PLC_TO_PC.DATA[79] := ' ';
   PLC_TO_PC.DATA[80] := ' ';
   PLC_TO_PC.DATA[81] := ' ';
   PLC_TO_PC.DATA[82] := ' ';
   PLC_TO_PC.DATA[83] := ' ';
   PLC_TO_PC.DATA[84] := ' ';
   PLC_TO_PC.DATA[85] := ' ';
   PLC_TO_PC.DATA[86] := ' ';
   PLC_TO_PC.DATA[87] := ' ';
   PLC_TO_PC.DATA[88] := ' ';
   PLC_TO_PC.DATA[89] := ' ';
   PLC_TO_PC.DATA[90] := ' ';
   PLC_TO_PC.DATA[91] := ' ';
   PLC_TO_PC.DATA[92] := ' ';
   PLC_TO_PC.DATA[93] := ' ';
   PLC_TO_PC.DATA[94] := ' ';
   PLC_TO_PC.DATA[95] := ' ';
   PLC_TO_PC.DATA[96] := ' ';
   PLC_TO_PC.DATA[97] := ' ';
   PLC_TO_PC.DATA[98] := ' ';
   PLC_TO_PC.DATA[99] := ' ';
   PLC_TO_PC.DATA[100] := ' ';
   PLC_TO_PC.DATA[101] := ' ';
   PLC_TO_PC.DATA[102] := ' ';
   PLC_TO_PC.DATA[103] := ' ';
   PLC_TO_PC.DATA[104] := ' ';
   PLC_TO_PC.DATA[105] := ' ';
   PLC_TO_PC.DATA[106] := ' ';
   PLC_TO_PC.DATA[107] := ' ';
   PLC_TO_PC.DATA[108] := ' ';
   PLC_TO_PC.DATA[109] := ' ';
   PLC_TO_PC.DATA[110] := ' ';
   PLC_TO_PC.DATA[111] := ' ';
   PLC_TO_PC.DATA[112] := ' ';
   PLC_TO_PC.DATA[113] := ' ';
   PLC_TO_PC.DATA[114] := ' ';
   PLC_TO_PC.DATA[115] := ' ';
   PLC_TO_PC.DATA[116] := ' ';
   PLC_TO_PC.DATA[117] := ' ';
   PLC_TO_PC.DATA[118] := ' ';
   PLC_TO_PC.DATA[119] := ' ';
   PLC_TO_PC.DATA[120] := ' ';
   PLC_TO_PC.DATA[121] := ' ';
   PLC_TO_PC.DATA[122] := ' ';
   PLC_TO_PC.DATA[123] := ' ';
   PLC_TO_PC.DATA[124] := ' ';
   PLC_TO_PC.DATA[125] := ' ';
   PLC_TO_PC.DATA[126] := ' ';
   PLC_TO_PC.DATA[127] := ' ';
   PLC_TO_PC.DATA[128] := ' ';
   PLC_TO_PC.DATA[129] := ' ';
   PLC_TO_PC.DATA[130] := ' ';
   PLC_TO_PC.DATA[131] := ' ';
   PLC_TO_PC.DATA[132] := ' ';
   PLC_TO_PC.DATA[133] := ' ';
   PLC_TO_PC.DATA[134] := ' ';
   PLC_TO_PC.DATA[135] := ' ';
   PLC_TO_PC.DATA[136] := ' ';
   PLC_TO_PC.DATA[137] := ' ';
   PLC_TO_PC.DATA[138] := ' ';
   PLC_TO_PC.DATA[139] := ' ';
   PLC_TO_PC.DATA[140] := ' ';
   PLC_TO_PC.DATA[141] := ' ';
   PLC_TO_PC.DATA[142] := ' ';
   PLC_TO_PC.DATA[143] := ' ';
   PLC_TO_PC.DATA[144] := ' ';
   PLC_TO_PC.DATA[145] := ' ';
   PLC_TO_PC.DATA[146] := ' ';
   PLC_TO_PC.DATA[147] := ' ';
   PLC_TO_PC.DATA[148] := ' ';
   PLC_TO_PC.DATA[149] := ' ';
   PLC_TO_PC.DATA[150] := ' ';
   PLC_TO_PC.DATA[151] := ' ';
   PLC_TO_PC.DATA[152] := ' ';
   PLC_TO_PC.DATA[153] := ' ';
   PLC_TO_PC.DATA[154] := ' ';
   PLC_TO_PC.DATA[155] := ' ';
   PLC_TO_PC.DATA[156] := ' ';
   PLC_TO_PC.DATA[157] := ' ';
   PLC_TO_PC.DATA[158] := ' ';
   PLC_TO_PC.DATA[159] := ' ';
   PLC_TO_PC.DATA[160] := ' ';
   PLC_TO_PC.DATA[161] := ' ';
   PLC_TO_PC.DATA[162] := ' ';
   PLC_TO_PC.DATA[163] := ' ';
   PLC_TO_PC.DATA[164] := ' ';
   PLC_TO_PC.DATA[165] := ' ';
   PLC_TO_PC.DATA[166] := ' ';
   PLC_TO_PC.DATA[167] := ' ';
   PLC_TO_PC.DATA[168] := ' ';
   PLC_TO_PC.DATA[169] := ' ';
   PLC_TO_PC.DATA[170] := ' ';
   PLC_TO_PC.DATA[171] := ' ';
   PLC_TO_PC.DATA[172] := ' ';
   PLC_TO_PC.DATA[173] := ' ';
   PLC_TO_PC.DATA[174] := ' ';
   PLC_TO_PC.DATA[175] := ' ';
   PLC_TO_PC.DATA[176] := ' ';
   PLC_TO_PC.DATA[177] := ' ';
   PLC_TO_PC.DATA[178] := ' ';
   PLC_TO_PC.DATA[179] := ' ';
   PLC_TO_PC.DATA[180] := ' ';
   PLC_TO_PC.DATA[181] := ' ';
   PLC_TO_PC.DATA[182] := ' ';
   PLC_TO_PC.DATA[183] := ' ';
   PLC_TO_PC.DATA[184] := ' ';
   PLC_TO_PC.DATA[185] := ' ';
   PLC_TO_PC.DATA[186] := ' ';
   PLC_TO_PC.DATA[187] := ' ';
   PLC_TO_PC.DATA[188] := ' ';
   PLC_TO_PC.DATA[189] := ' ';
   PLC_TO_PC.DATA[190] := ' ';
   PLC_TO_PC.DATA[191] := ' ';
   PLC_TO_PC.DATA[192] := ' ';
   PLC_TO_PC.DATA[193] := ' ';
   PLC_TO_PC.DATA[194] := ' ';
   PLC_TO_PC.DATA[195] := ' ';
   PLC_TO_PC.DATA[196] := ' ';
   PLC_TO_PC.DATA[197] := ' ';
   PLC_TO_PC.DATA[198] := ' ';
   PLC_TO_PC.DATA[199] := ' ';
   PLC_TO_PC.DATA[200] := ' ';
   PLC_TO_PC.DATA[201] := ' ';
   PLC_TO_PC.DATA[202] := ' ';
   PLC_TO_PC.DATA[203] := ' ';
   PLC_TO_PC.DATA[204] := ' ';
   PLC_TO_PC.DATA[205] := ' ';
   PLC_TO_PC.DATA[206] := ' ';
   PLC_TO_PC.DATA[207] := ' ';
   PLC_TO_PC.DATA[208] := ' ';
   PLC_TO_PC.DATA[209] := ' ';
   PLC_TO_PC.DATA[210] := ' ';
   PLC_TO_PC.DATA[211] := ' ';
   PLC_TO_PC.DATA[212] := ' ';
   PLC_TO_PC.DATA[213] := ' ';
   PLC_TO_PC.DATA[214] := ' ';
   PLC_TO_PC.DATA[215] := ' ';
   PLC_TO_PC.DATA[216] := ' ';
   PLC_TO_PC.DATA[217] := ' ';
   PLC_TO_PC.DATA[218] := ' ';
   PLC_TO_PC.DATA[219] := ' ';
   PLC_TO_PC.DATA[220] := ' ';
   PLC_TO_PC.DATA[221] := ' ';
   PLC_TO_PC.DATA[222] := ' ';
   PLC_TO_PC.DATA[223] := ' ';
   PLC_TO_PC.DATA[224] := ' ';
   PLC_TO_PC.DATA[225] := ' ';
   PLC_TO_PC.DATA[226] := ' ';
   PLC_TO_PC.DATA[227] := ' ';
   PLC_TO_PC.DATA[228] := ' ';
   PLC_TO_PC.DATA[229] := ' ';
   PLC_TO_PC.DATA[230] := ' ';
   PLC_TO_PC.DATA[231] := ' ';
   PLC_TO_PC.DATA[232] := ' ';
   PLC_TO_PC.DATA[233] := ' ';
   PLC_TO_PC.DATA[234] := ' ';
   PLC_TO_PC.DATA[235] := ' ';
   PLC_TO_PC.DATA[236] := ' ';
   PLC_TO_PC.DATA[237] := ' ';
   PLC_TO_PC.DATA[238] := ' ';
   PLC_TO_PC.DATA[239] := ' ';
   PLC_TO_PC.DATA[240] := ' ';
   PLC_TO_PC.DATA[241] := ' ';
   PLC_TO_PC.DATA[242] := ' ';
   PLC_TO_PC.DATA[243] := ' ';
   PLC_TO_PC.DATA[244] := ' ';
   PLC_TO_PC.DATA[245] := ' ';
   PLC_TO_PC.DATA[246] := ' ';
   PLC_TO_PC.DATA[247] := ' ';
   PLC_TO_PC.DATA[248] := ' ';
   PLC_TO_PC.DATA[249] := ' ';
   PLC_TO_PC.DATA[250] := ' ';
   PLC_TO_PC.DATA[251] := ' ';
   PLC_TO_PC.DATA[252] := ' ';
   PLC_TO_PC.DATA[253] := ' ';
   PLC_TO_PC.DATA[254] := ' ';
   PLC_TO_PC.DATA[255] := ' ';
   PLC_TO_PC.DATA[256] := ' ';
   PLC_TO_PC.DATA[257] := ' ';
   PLC_TO_PC.DATA[258] := ' ';
   PLC_TO_PC.DATA[259] := ' ';
   PLC_TO_PC.DATA[260] := ' ';
   PLC_TO_PC.DATA[261] := ' ';
   PLC_TO_PC.DATA[262] := ' ';
   PLC_TO_PC.DATA[263] := ' ';
   PLC_TO_PC.DATA[264] := ' ';
   PLC_TO_PC.DATA[265] := ' ';
   PLC_TO_PC.DATA[266] := ' ';
   PLC_TO_PC.DATA[267] := ' ';
   PLC_TO_PC.DATA[268] := ' ';
   PLC_TO_PC.DATA[269] := ' ';
   PLC_TO_PC.DATA[270] := ' ';
   PLC_TO_PC.DATA[271] := ' ';
   PLC_TO_PC.DATA[272] := ' ';
   PLC_TO_PC.DATA[273] := ' ';
   PLC_TO_PC.DATA[274] := ' ';
   PLC_TO_PC.DATA[275] := ' ';
   PLC_TO_PC.DATA[276] := ' ';
   PLC_TO_PC.DATA[277] := ' ';
   PLC_TO_PC.DATA[278] := ' ';
   PLC_TO_PC.DATA[279] := ' ';
   PLC_TO_PC.DATA[280] := ' ';
   PLC_TO_PC.DATA[281] := ' ';
   PLC_TO_PC.DATA[282] := ' ';
   PLC_TO_PC.DATA[283] := ' ';
   PLC_TO_PC.DATA[284] := ' ';
   PLC_TO_PC.DATA[285] := ' ';
   PLC_TO_PC.DATA[286] := ' ';
   PLC_TO_PC.DATA[287] := ' ';
   PLC_TO_PC.DATA[288] := ' ';
   PLC_TO_PC.DATA[289] := ' ';
   PLC_TO_PC.DATA[290] := ' ';
   PLC_TO_PC.DATA[291] := ' ';
   PLC_TO_PC.DATA[292] := ' ';
   PLC_TO_PC.DATA[293] := ' ';
   PLC_TO_PC.DATA[294] := ' ';
   PLC_TO_PC.DATA[295] := ' ';
   PLC_TO_PC.DATA[296] := ' ';
   PLC_TO_PC.DATA[297] := ' ';
   PLC_TO_PC.DATA[298] := ' ';
   PLC_TO_PC.DATA[299] := ' ';
   PLC_TO_PC.DATA[300] := ' ';
   PLC_TO_PC.DATA[301] := ' ';
   PLC_TO_PC.DATA[302] := ' ';
   PLC_TO_PC.DATA[303] := ' ';
   PLC_TO_PC.DATA[304] := ' ';
   PLC_TO_PC.DATA[305] := ' ';
   PLC_TO_PC.DATA[306] := ' ';
   PLC_TO_PC.DATA[307] := ' ';
   PLC_TO_PC.DATA[308] := ' ';
   PLC_TO_PC.DATA[309] := ' ';
   PLC_TO_PC.DATA[310] := ' ';
   PLC_TO_PC.DATA[311] := ' ';
   PLC_TO_PC.DATA[312] := ' ';
   PLC_TO_PC.DATA[313] := ' ';
   PLC_TO_PC.DATA[314] := ' ';
   PLC_TO_PC.DATA[315] := ' ';
   PLC_TO_PC.DATA[316] := ' ';
   PLC_TO_PC.DATA[317] := ' ';
   PLC_TO_PC.DATA[318] := ' ';
   PLC_TO_PC.DATA[319] := ' ';
   PLC_TO_PC.DATA[320] := ' ';
   PLC_TO_PC.DATA[321] := ' ';
   PLC_TO_PC.DATA[322] := ' ';
   PLC_TO_PC.DATA[323] := ' ';